(* Logix 5000 project; controller MV vendor 1 type 14 code 217 rev 31.11; software revision 31.00; part 26 of 53 *)
(* tags used below, declared in another part *)
   CWD : CHECKWORD_FLAGS;
   IGI_TestBit : BOOL;
   MC_B12 : INT[255];   // PX SWITCH Proxy switch flags f ile
   MC_B3 : INT[255];   // BINARY
   MC_COMMS_FROM_BLUNGER : MESSAGE;
   MC_COMMS_FROM_FV_ROUTING_PLC : MESSAGE;
   MC_COMMS_FROM_MV_ROUTING_PLC : MESSAGE;
   MC_N100 : INT[255];   // C1_PLC Channel 1 PLC data
   MC_N112 : INT[255];   // FVR DATA Data read from FV ro uting PLC
   MC_N113 : INT[255];   // MVR DATA Data read from MV ro uting PLC
   MC_N114 : INT[255];   // YP DATA
   MC_N120 : INT[255];   // C2 PLC Channel 2 PLC data
   MC_R2_SW1 : PlantItem;   // R2_SW1
   MC_R2_SW2 : PlantItem;   // R2_SW2
   MC_R2_SW3 : PlantItem;   // R2_SW3
   MC_R2_SW3_1 : PlantItem;   // R2_SW3_1
   MC_R2_SW4 : PlantItem;   // R2_SW4
   MC_R3_SW1 : PlantItem;   // R3_SW1
   MC_R3_SW2 : PlantItem;   // R3_SW2
   MC_R3_SW2_1 : PlantItem;   // PROXY
   MC_R4_SW1 : PlantItem;   // R4_SW1
   MC_R4_SW2 : PlantItem;   // R4_SW2
   MC_R4_SW3 : PlantItem;   // R4_SW3
   MC_R4_SW4 : PlantItem;   // R4_SW4
   MC_R4_SW6 : PlantItem;   // R4_SW6
   MC_R6_SW1 : PlantItem;   // R6_SW1
   MC_T4 : TIMER[255];   // TIMER
(* MC_Common, continued *)

ROUTINE MC_PX_SWITCH_12   (* ladder *)
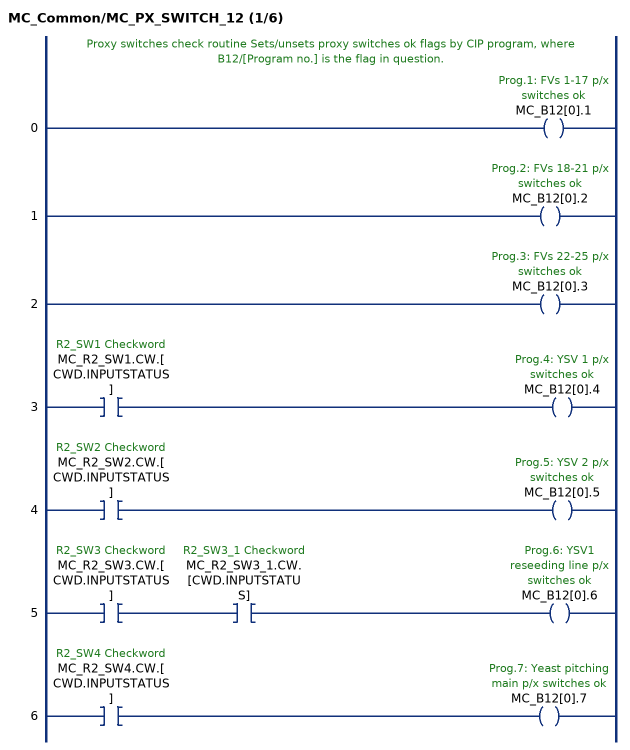
   // Proxy switches check routine Sets/unsets proxy switches ok flags by CIP program, where B12/[Program no.] is the flag in question.
   0: OTE(MC_B12[0].1);
   1: OTE(MC_B12[0].2);
   2: OTE(MC_B12[0].3);
   3: XIC(MC_R2_SW1.CW.[CWD.INPUTSTATUS])OTE(MC_B12[0].4);
   4: XIC(MC_R2_SW2.CW.[CWD.INPUTSTATUS])OTE(MC_B12[0].5);
   5: XIC(MC_R2_SW3.CW.[CWD.INPUTSTATUS])XIC(MC_R2_SW3_1.CW.[CWD.INPUTSTATUS])OTE(MC_B12[0].6);
   6: XIC(MC_R2_SW4.CW.[CWD.INPUTSTATUS])OTE(MC_B12[0].7);
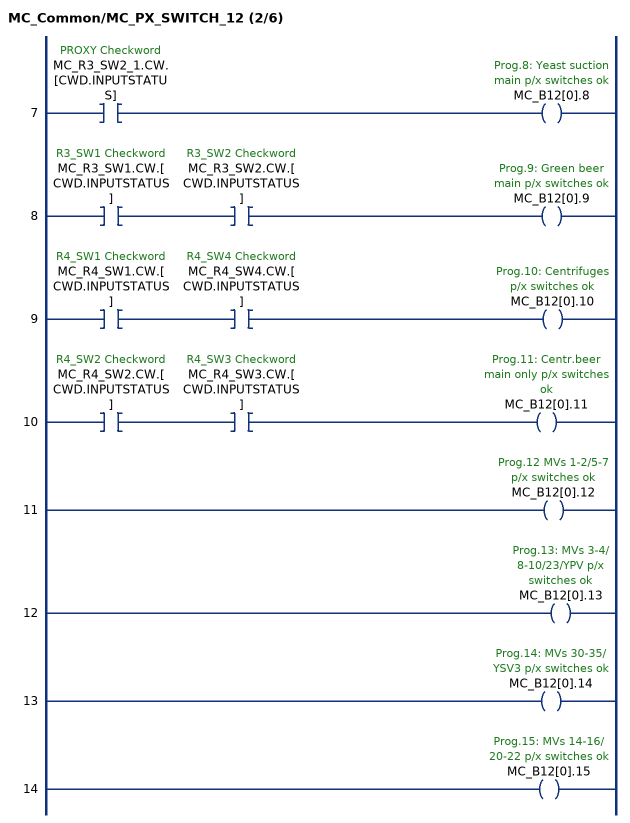
   7: XIC(MC_R3_SW2_1.CW.[CWD.INPUTSTATUS])OTE(MC_B12[0].8);
   8: XIC(MC_R3_SW1.CW.[CWD.INPUTSTATUS])XIC(MC_R3_SW2.CW.[CWD.INPUTSTATUS])OTE(MC_B12[0].9);
   9: XIC(MC_R4_SW1.CW.[CWD.INPUTSTATUS])XIC(MC_R4_SW4.CW.[CWD.INPUTSTATUS])OTE(MC_B12[0].10);
   10: XIC(MC_R4_SW2.CW.[CWD.INPUTSTATUS])XIC(MC_R4_SW3.CW.[CWD.INPUTSTATUS])OTE(MC_B12[0].11);
   11: OTE(MC_B12[0].12);
   12: OTE(MC_B12[0].13);
   13: OTE(MC_B12[0].14);
   14: OTE(MC_B12[0].15);
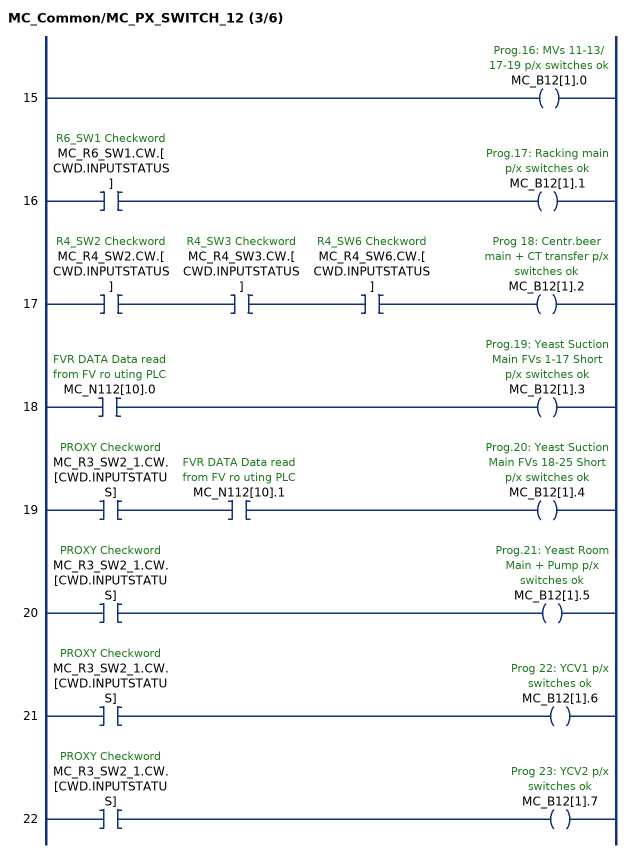
   15: OTE(MC_B12[1].0);
   16: XIC(MC_R6_SW1.CW.[CWD.INPUTSTATUS])OTE(MC_B12[1].1);
   17: XIC(MC_R4_SW2.CW.[CWD.INPUTSTATUS])XIC(MC_R4_SW3.CW.[CWD.INPUTSTATUS])XIC(MC_R4_SW6.CW.[CWD.INPUTSTATUS])OTE(MC_B12[1].2);
   18: XIC(MC_N112[10].0)OTE(MC_B12[1].3);
   19: XIC(MC_R3_SW2_1.CW.[CWD.INPUTSTATUS])XIC(MC_N112[10].1)OTE(MC_B12[1].4);
   20: XIC(MC_R3_SW2_1.CW.[CWD.INPUTSTATUS])OTE(MC_B12[1].5);
   21: XIC(MC_R3_SW2_1.CW.[CWD.INPUTSTATUS])OTE(MC_B12[1].6);
   22: XIC(MC_R3_SW2_1.CW.[CWD.INPUTSTATUS])OTE(MC_B12[1].7);
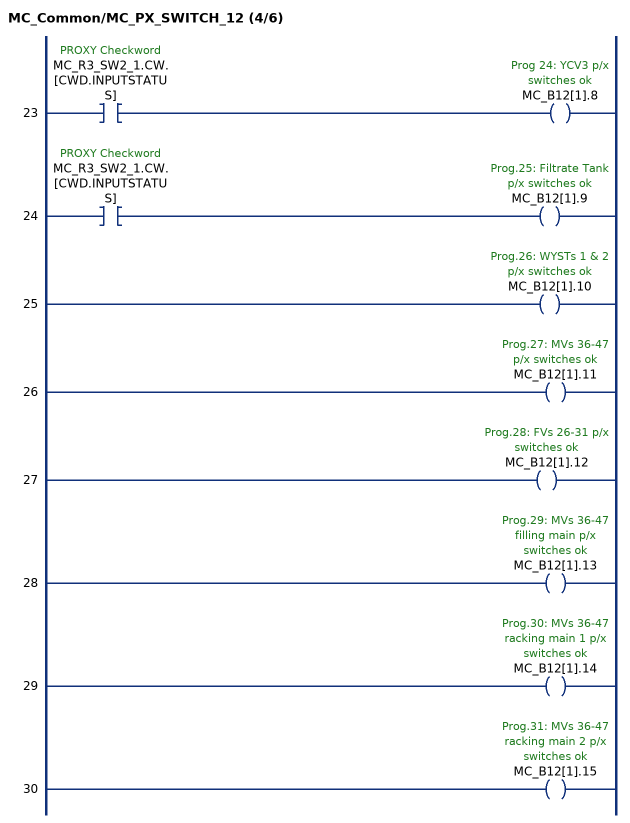
   23: XIC(MC_R3_SW2_1.CW.[CWD.INPUTSTATUS])OTE(MC_B12[1].8);
   24: XIC(MC_R3_SW2_1.CW.[CWD.INPUTSTATUS])OTE(MC_B12[1].9);
   25: OTE(MC_B12[1].10);
   26: OTE(MC_B12[1].11);
   27: OTE(MC_B12[1].12);
   28: OTE(MC_B12[1].13);
   29: OTE(MC_B12[1].14);
   30: OTE(MC_B12[1].15);
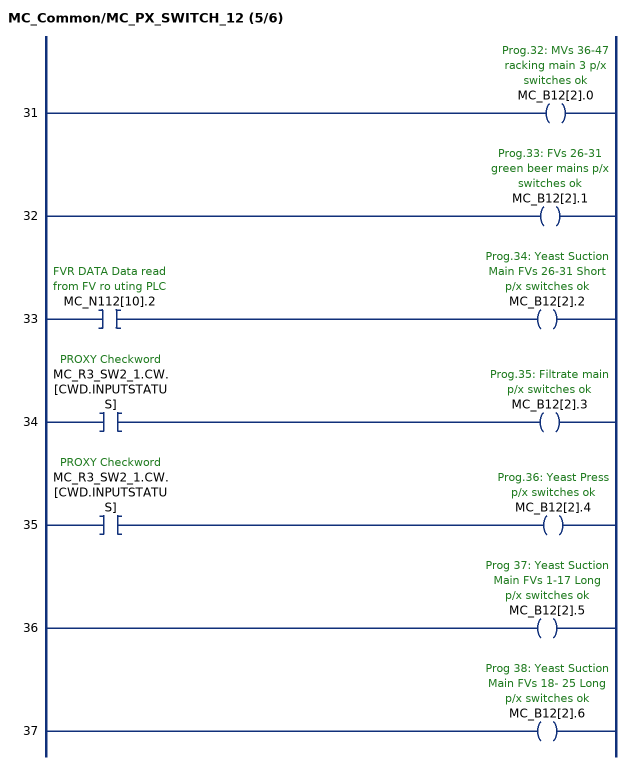
   31: OTE(MC_B12[2].0);
   32: OTE(MC_B12[2].1);
   33: XIC(MC_N112[10].2)OTE(MC_B12[2].2);
   34: XIC(MC_R3_SW2_1.CW.[CWD.INPUTSTATUS])OTE(MC_B12[2].3);
   35: XIC(MC_R3_SW2_1.CW.[CWD.INPUTSTATUS])OTE(MC_B12[2].4);
   36: OTE(MC_B12[2].5);
   37: OTE(MC_B12[2].6);
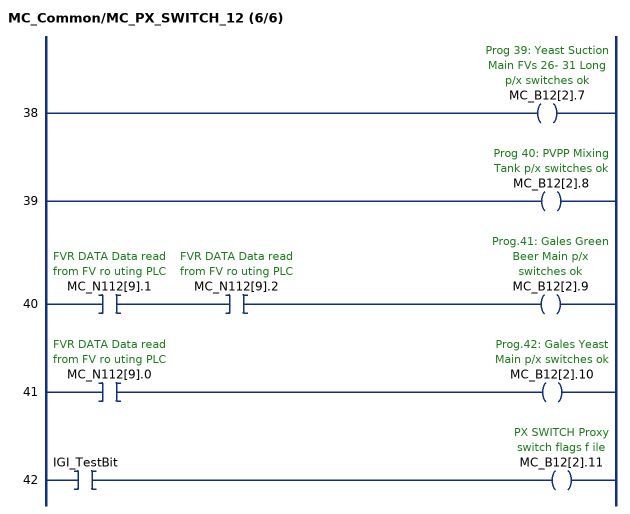
   38: OTE(MC_B12[2].7);
   39: OTE(MC_B12[2].8);
   40: XIC(MC_N112[9].1)XIC(MC_N112[9].2)OTE(MC_B12[2].9);
   41: XIC(MC_N112[9].0)OTE(MC_B12[2].10);
   42: XIC(IGI_TestBit)OTE(MC_B12[2].11);
END_ROUTINE

ROUTINE MC_REMOTE_SYS_245   (* ladder *)
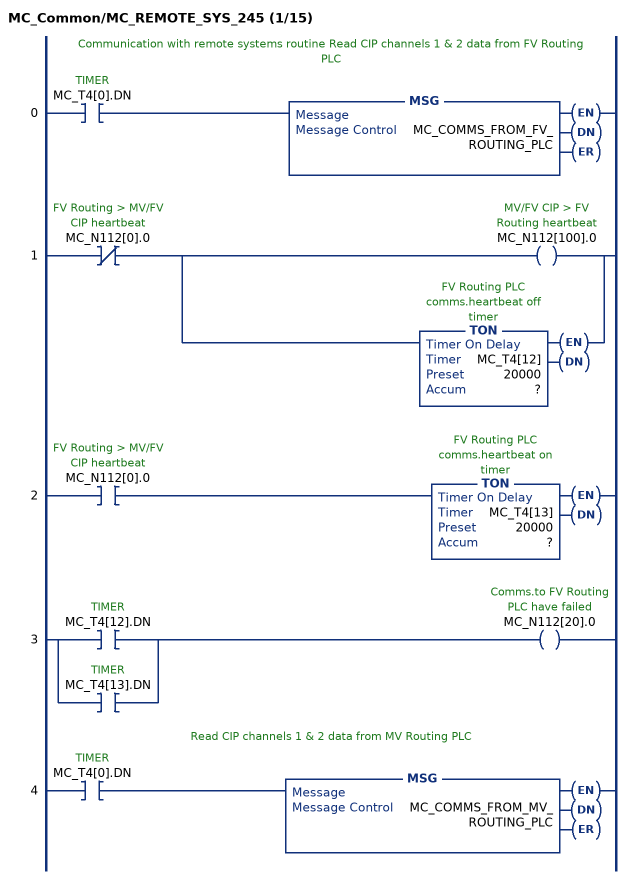
   // Communication with remote systems routine Read CIP channels 1 & 2 data from FV Routing PLC
   0: XIC(MC_T4[0].DN)MSG(MC_COMMS_FROM_FV_ROUTING_PLC);
   1: XIO(MC_N112[0].0)[OTE(MC_N112[100].0) ,TON(MC_T4[12],?,?) ];
   2: XIC(MC_N112[0].0)TON(MC_T4[13],?,?);
   3: [XIC(MC_T4[12].DN) ,XIC(MC_T4[13].DN) ]OTE(MC_N112[20].0);
   // Read CIP channels 1 & 2 data from MV Routing PLC
   4: XIC(MC_T4[0].DN)MSG(MC_COMMS_FROM_MV_ROUTING_PLC);
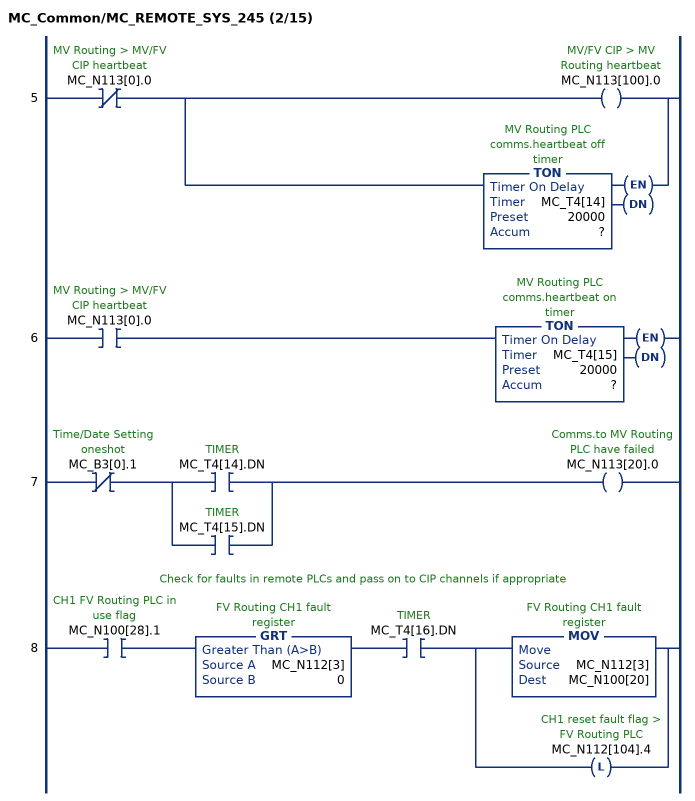
   5: XIO(MC_N113[0].0)[OTE(MC_N113[100].0) ,TON(MC_T4[14],?,?) ];
   6: XIC(MC_N113[0].0)TON(MC_T4[15],?,?);
   7: XIO(MC_B3[0].1)[XIC(MC_T4[14].DN) ,XIC(MC_T4[15].DN) ]OTE(MC_N113[20].0);
   // Check for faults in remote PLCs and pass on to CIP channels if appropriate
   8: XIC(MC_N100[28].1)GRT(MC_N112[3],0)XIC(MC_T4[16].DN)[MOV(MC_N112[3],MC_N100[20]) ,OTL(MC_N112[104].4) ];
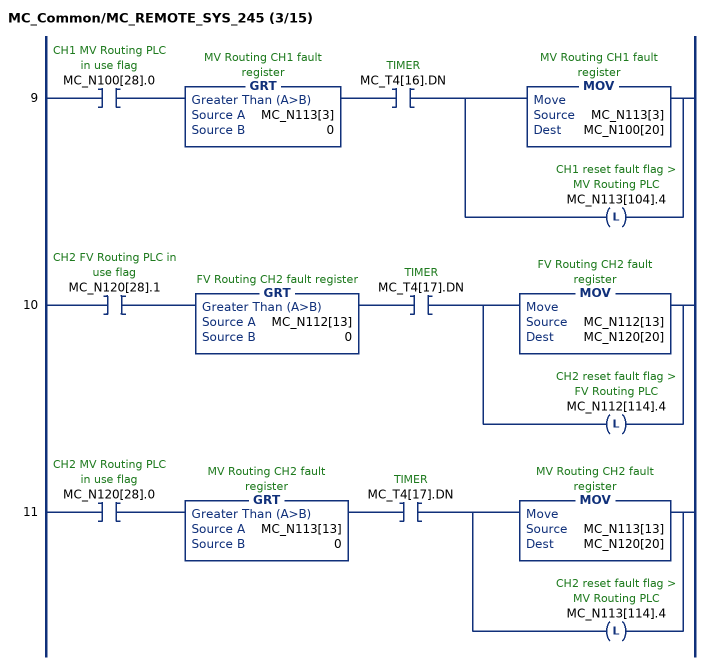
   9: XIC(MC_N100[28].0)GRT(MC_N113[3],0)XIC(MC_T4[16].DN)[MOV(MC_N113[3],MC_N100[20]) ,OTL(MC_N113[104].4) ];
   10: XIC(MC_N120[28].1)GRT(MC_N112[13],0)XIC(MC_T4[17].DN)[MOV(MC_N112[13],MC_N120[20]) ,OTL(MC_N112[114].4) ];
   11: XIC(MC_N120[28].0)GRT(MC_N113[13],0)XIC(MC_T4[17].DN)[MOV(MC_N113[13],MC_N120[20]) ,OTL(MC_N113[114].4) ];
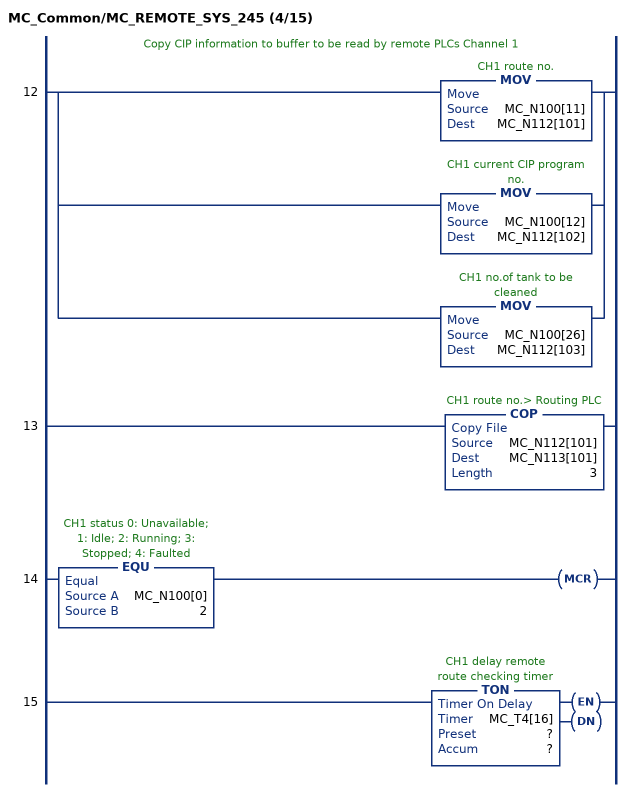
   // Copy CIP information to buffer to be read by remote PLCs Channel 1
   12: [MOV(MC_N100[11],MC_N112[101]) ,MOV(MC_N100[12],MC_N112[102]) ,MOV(MC_N100[26],MC_N112[103]) ];
   13: COP(MC_N112[101],MC_N113[101],3);
   14: EQU(MC_N100[0],2)MCR();
   15: TON(MC_T4[16],?,?);
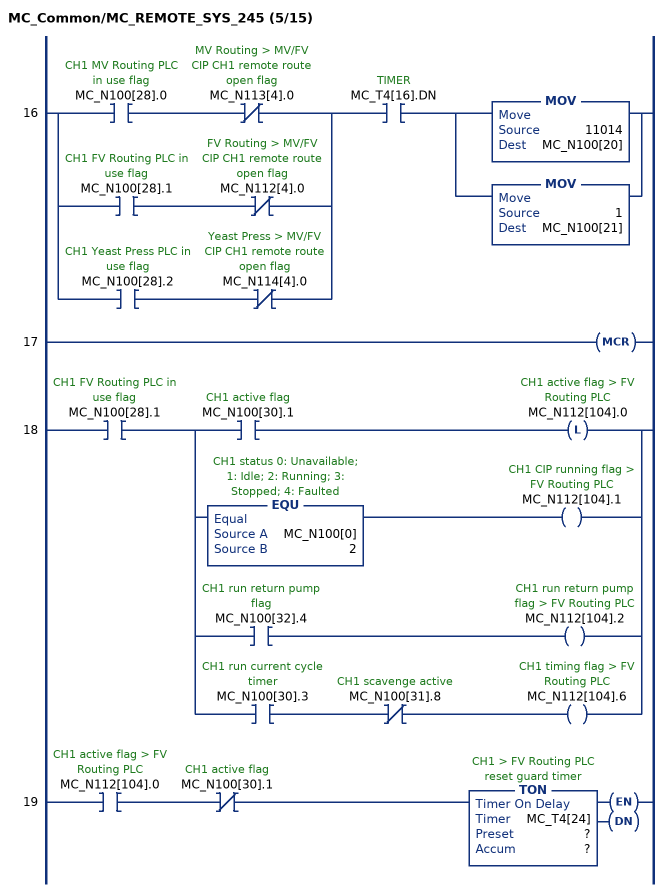
   16: [XIC(MC_N100[28].0) XIO(MC_N113[4].0) ,XIC(MC_N100[28].1) XIO(MC_N112[4].0) ,XIC(MC_N100[28].2) XIO(MC_N114[4].0) ]XIC(MC_T4[16].DN)[MOV(11014,MC_N100[20]) ,MOV(1,MC_N100[21]) ];
   17: MCR();
   18: XIC(MC_N100[28].1)[XIC(MC_N100[30].1) OTL(MC_N112[104].0) ,EQU(MC_N100[0],2) OTE(MC_N112[104].1) ,XIC(MC_N100[32].4) OTE(MC_N112[104].2) ,XIC(MC_N100[30].3) XIO(MC_N100[31].8) OTE(MC_N112[104].6) ];
   19: XIC(MC_N112[104].0)XIO(MC_N100[30].1)TON(MC_T4[24],?,?);
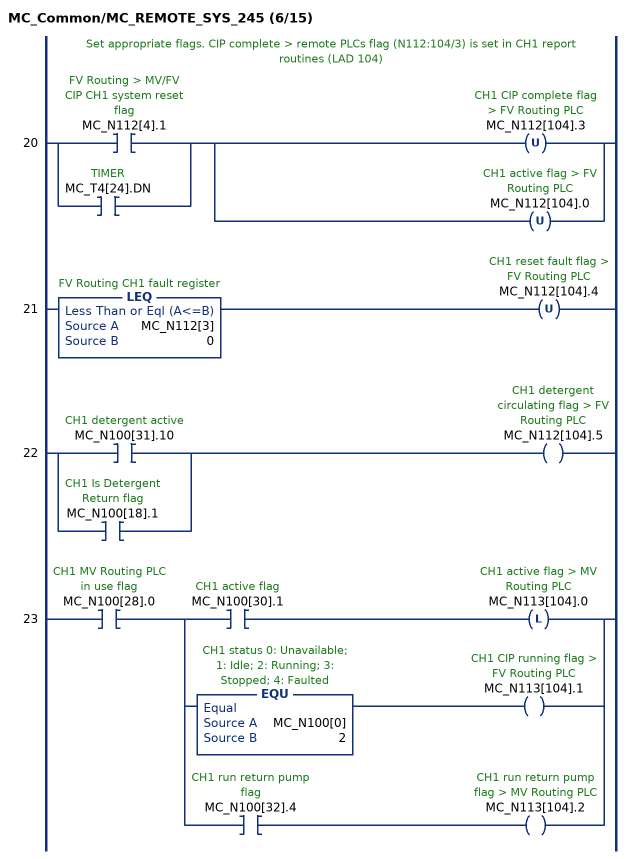
   // Set appropriate flags. CIP complete > remote PLCs flag (N112:104/3) is set in CH1 report routines (LAD 104)
   20: [XIC(MC_N112[4].1) ,XIC(MC_T4[24].DN) ][OTU(MC_N112[104].3) ,OTU(MC_N112[104].0) ];
   21: LEQ(MC_N112[3],0)OTU(MC_N112[104].4);
   22: [XIC(MC_N100[31].10) ,XIC(MC_N100[18].1) ]OTE(MC_N112[104].5);
   23: XIC(MC_N100[28].0)[XIC(MC_N100[30].1) OTL(MC_N113[104].0) ,EQU(MC_N100[0],2) OTE(MC_N113[104].1) ,XIC(MC_N100[32].4) OTE(MC_N113[104].2) ];
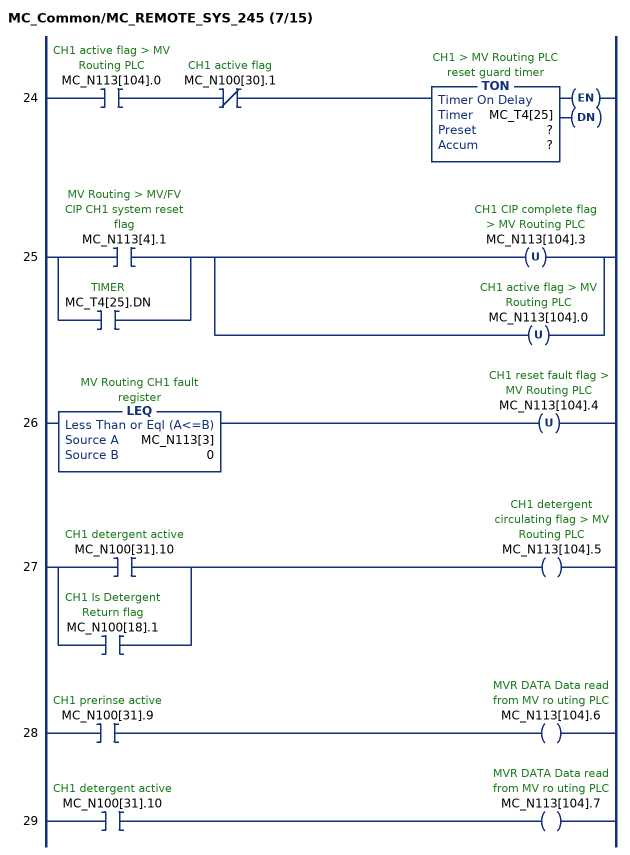
   24: XIC(MC_N113[104].0)XIO(MC_N100[30].1)TON(MC_T4[25],?,?);
   25: [XIC(MC_N113[4].1) ,XIC(MC_T4[25].DN) ][OTU(MC_N113[104].3) ,OTU(MC_N113[104].0) ];
   26: LEQ(MC_N113[3],0)OTU(MC_N113[104].4);
   27: [XIC(MC_N100[31].10) ,XIC(MC_N100[18].1) ]OTE(MC_N113[104].5);
   28: XIC(MC_N100[31].9)OTE(MC_N113[104].6);
   29: XIC(MC_N100[31].10)OTE(MC_N113[104].7);
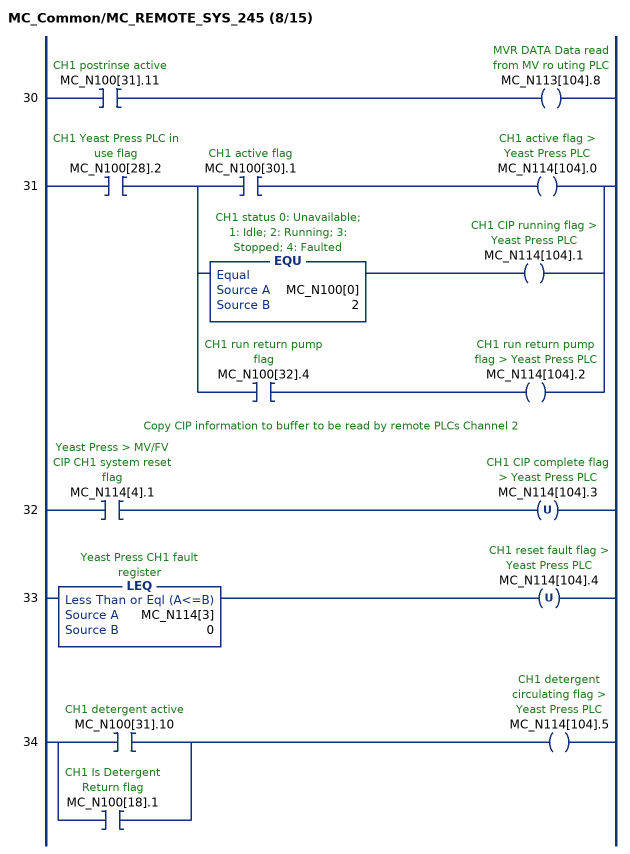
   30: XIC(MC_N100[31].11)OTE(MC_N113[104].8);
   31: XIC(MC_N100[28].2)[XIC(MC_N100[30].1) OTE(MC_N114[104].0) ,EQU(MC_N100[0],2) OTE(MC_N114[104].1) ,XIC(MC_N100[32].4) OTE(MC_N114[104].2) ];
   // Copy CIP information to buffer to be read by remote PLCs Channel 2
   32: XIC(MC_N114[4].1)OTU(MC_N114[104].3);
   33: LEQ(MC_N114[3],0)OTU(MC_N114[104].4);
   34: [XIC(MC_N100[31].10) ,XIC(MC_N100[18].1) ]OTE(MC_N114[104].5);
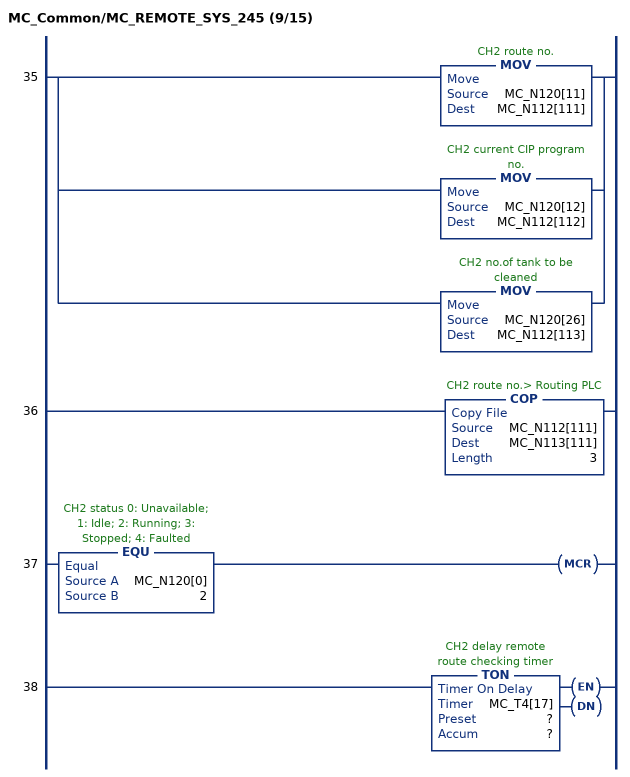
   35: [MOV(MC_N120[11],MC_N112[111]) ,MOV(MC_N120[12],MC_N112[112]) ,MOV(MC_N120[26],MC_N112[113]) ];
   36: COP(MC_N112[111],MC_N113[111],3);
   37: EQU(MC_N120[0],2)MCR();
   38: TON(MC_T4[17],?,?);
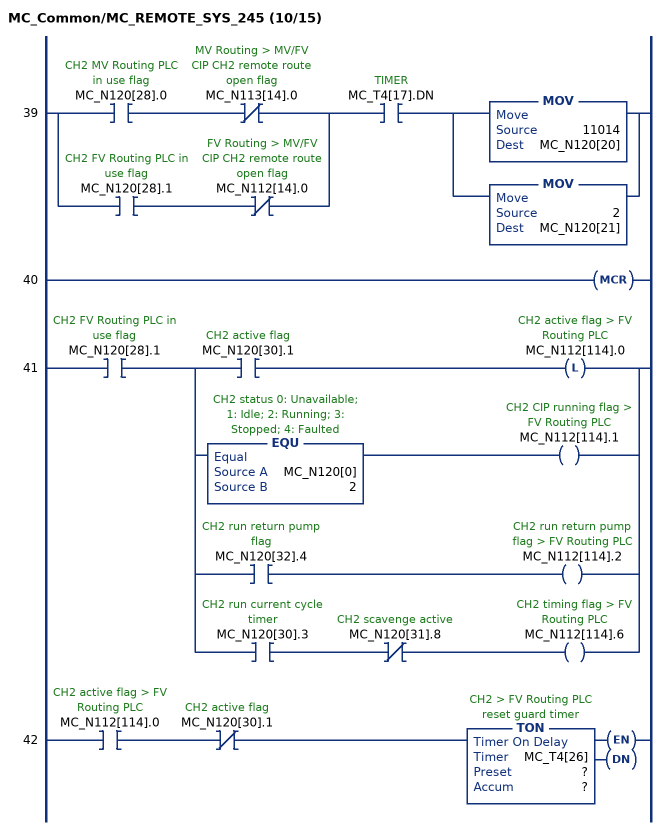
   39: [XIC(MC_N120[28].0) XIO(MC_N113[14].0) ,XIC(MC_N120[28].1) XIO(MC_N112[14].0) ]XIC(MC_T4[17].DN)[MOV(11014,MC_N120[20]) ,MOV(2,MC_N120[21]) ];
   40: MCR();
   41: XIC(MC_N120[28].1)[XIC(MC_N120[30].1) OTL(MC_N112[114].0) ,EQU(MC_N120[0],2) OTE(MC_N112[114].1) ,XIC(MC_N120[32].4) OTE(MC_N112[114].2) ,XIC(MC_N120[30].3) XIO(MC_N120[31].8) OTE(MC_N112[114].6) ];
   42: XIC(MC_N112[114].0)XIO(MC_N120[30].1)TON(MC_T4[26],?,?);
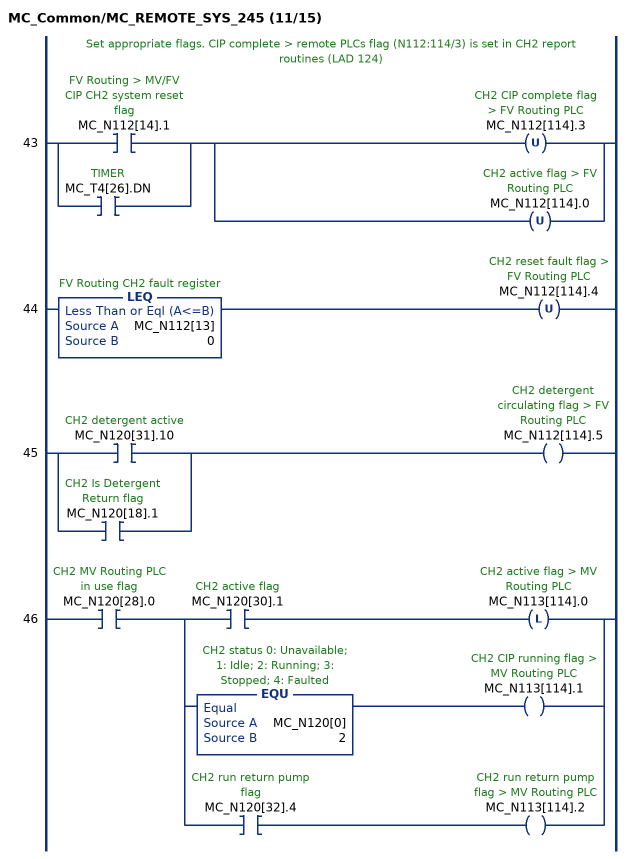
   // Set appropriate flags. CIP complete > remote PLCs flag (N112:114/3) is set in CH2 report routines (LAD 124)
   43: [XIC(MC_N112[14].1) ,XIC(MC_T4[26].DN) ][OTU(MC_N112[114].3) ,OTU(MC_N112[114].0) ];
   44: LEQ(MC_N112[13],0)OTU(MC_N112[114].4);
   45: [XIC(MC_N120[31].10) ,XIC(MC_N120[18].1) ]OTE(MC_N112[114].5);
   46: XIC(MC_N120[28].0)[XIC(MC_N120[30].1) OTL(MC_N113[114].0) ,EQU(MC_N120[0],2) OTE(MC_N113[114].1) ,XIC(MC_N120[32].4) OTE(MC_N113[114].2) ];
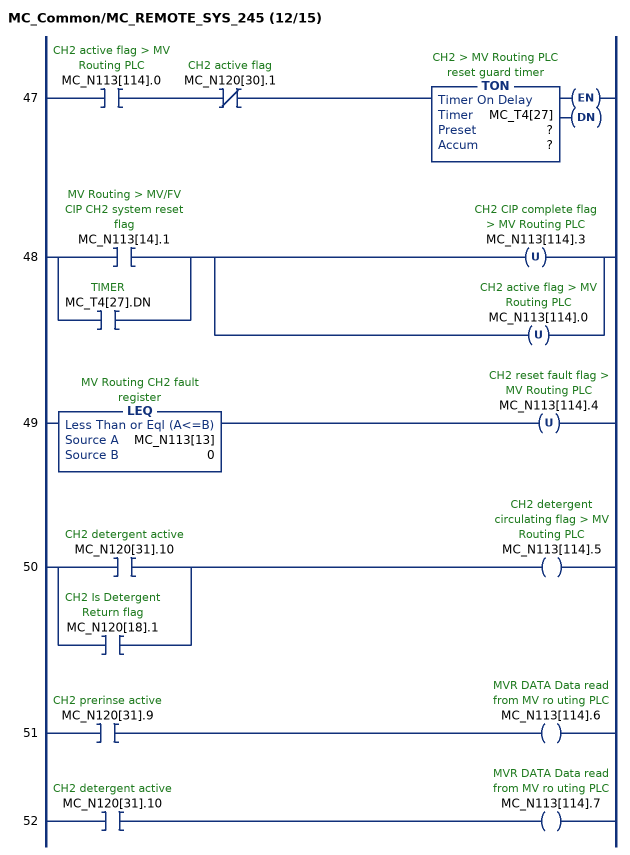
   47: XIC(MC_N113[114].0)XIO(MC_N120[30].1)TON(MC_T4[27],?,?);
   48: [XIC(MC_N113[14].1) ,XIC(MC_T4[27].DN) ][OTU(MC_N113[114].3) ,OTU(MC_N113[114].0) ];
   49: LEQ(MC_N113[13],0)OTU(MC_N113[114].4);
   50: [XIC(MC_N120[31].10) ,XIC(MC_N120[18].1) ]OTE(MC_N113[114].5);
   51: XIC(MC_N120[31].9)OTE(MC_N113[114].6);
   52: XIC(MC_N120[31].10)OTE(MC_N113[114].7);
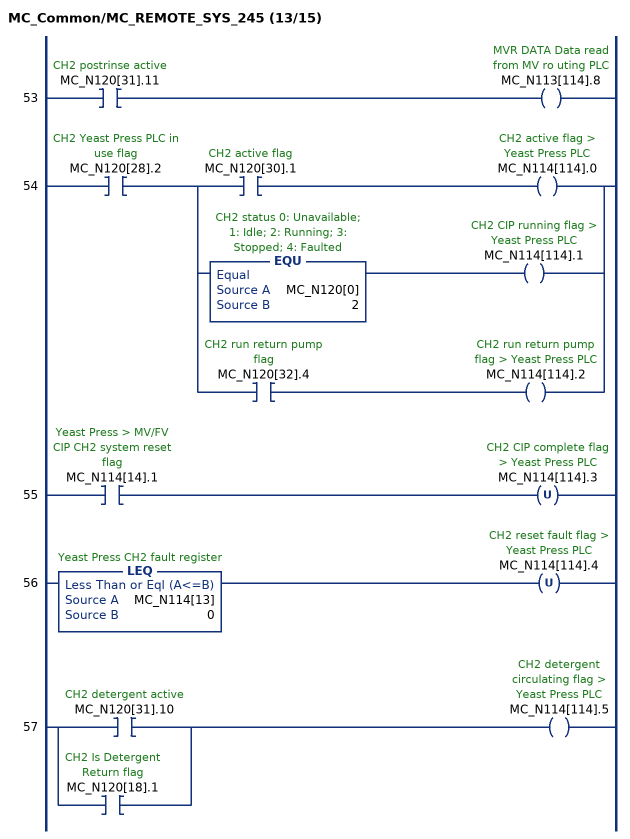
   53: XIC(MC_N120[31].11)OTE(MC_N113[114].8);
   54: XIC(MC_N120[28].2)[XIC(MC_N120[30].1) OTE(MC_N114[114].0) ,EQU(MC_N120[0],2) OTE(MC_N114[114].1) ,XIC(MC_N120[32].4) OTE(MC_N114[114].2) ];
   55: XIC(MC_N114[14].1)OTU(MC_N114[114].3);
   56: LEQ(MC_N114[13],0)OTU(MC_N114[114].4);
   57: [XIC(MC_N120[31].10) ,XIC(MC_N120[18].1) ]OTE(MC_N114[114].5);
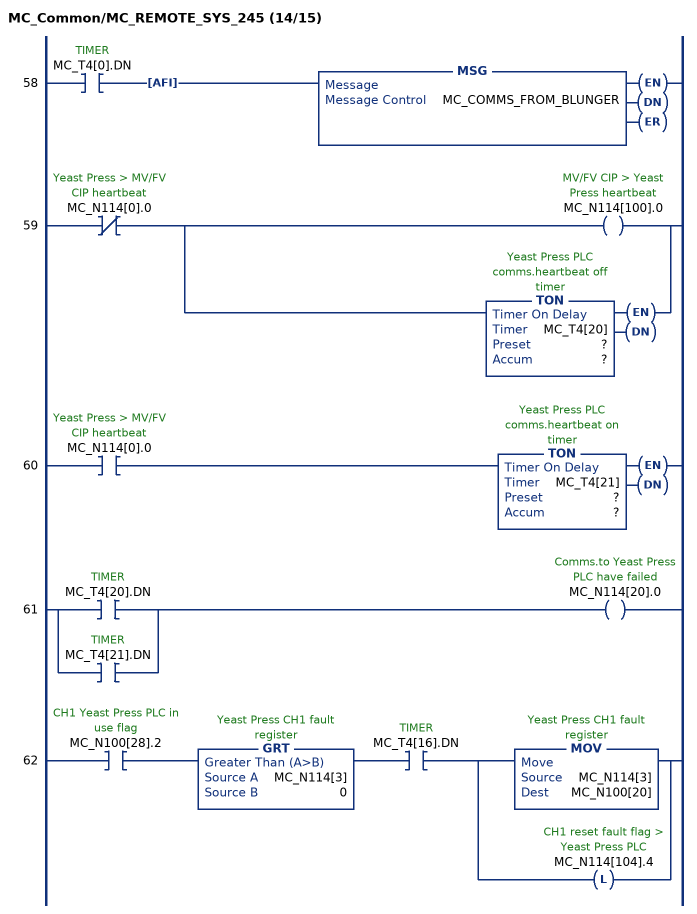
   58: XIC(MC_T4[0].DN)AFI()MSG(MC_COMMS_FROM_BLUNGER);
   59: XIO(MC_N114[0].0)[OTE(MC_N114[100].0) ,TON(MC_T4[20],?,?) ];
   60: XIC(MC_N114[0].0)TON(MC_T4[21],?,?);
   61: [XIC(MC_T4[20].DN) ,XIC(MC_T4[21].DN) ]OTE(MC_N114[20].0);
   62: XIC(MC_N100[28].2)GRT(MC_N114[3],0)XIC(MC_T4[16].DN)[MOV(MC_N114[3],MC_N100[20]) ,OTL(MC_N114[104].4) ];
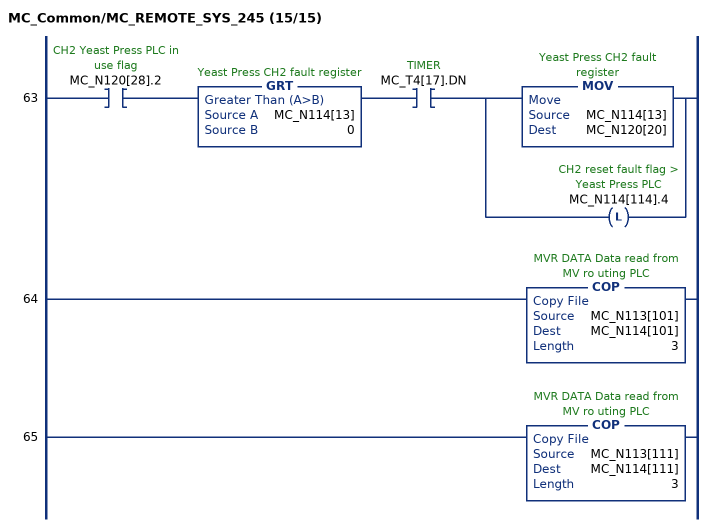
   63: XIC(MC_N120[28].2)GRT(MC_N114[13],0)XIC(MC_T4[17].DN)[MOV(MC_N114[13],MC_N120[20]) ,OTL(MC_N114[114].4) ];
   64: COP(MC_N113[101],MC_N114[101],3);
   65: COP(MC_N113[111],MC_N114[111],3);
END_ROUTINE
